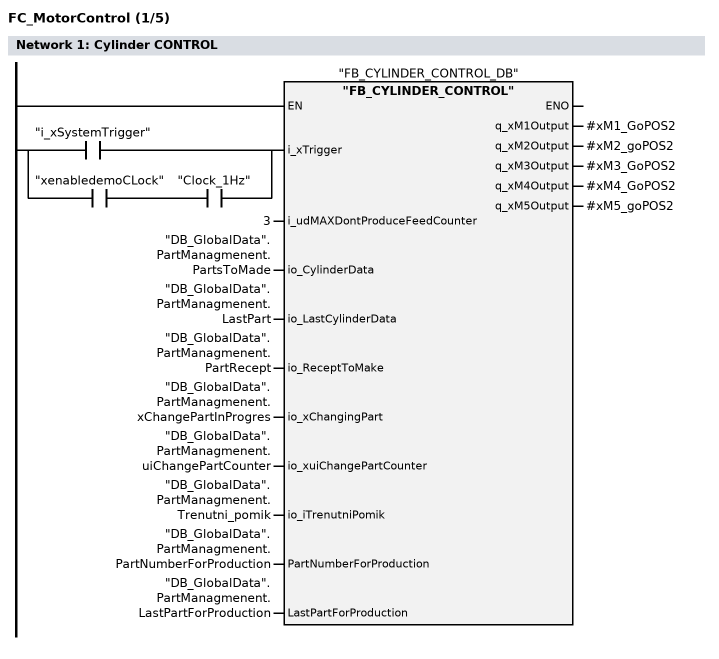
   RUNG wire#powerrail
      "FB_CYLINDER_CONTROL_DB"(i_xTrigger := wire#w1, i_udMAXDontProduceFeedCounter := 3, io_CylinderData := "DB_GlobalData".PartManagmenent.PartsToMade, io_LastCylinderData := "DB_GlobalData".PartManagmenent.LastPart, io_ReceptToMake := "DB_GlobalData".PartManagmenent.PartRecept, io_xChangingPart := "DB_GlobalData".PartManagmenent.xChangePartInProgres, io_xuiChangePartCounter := "DB_GlobalData".PartManagmenent.uiChangePartCounter, io_iTrenutniPomik := "DB_GlobalData".PartManagmenent.Trenutni_pomik, PartNumberForProduction := "DB_GlobalData".PartManagmenent.PartNumberForProduction, LastPartForProduction := "DB_GlobalData".PartManagmenent.LastPartForProduction, q_xM1Output => #xM1_GoPOS2, q_xM2Output => #xM2_goPOS2, q_xM3Output => #xM3_GoPOS2, q_xM4Output => #xM4_GoPOS2, q_xM5Output => #xM5_goPOS2)
   END_RUNG
   RUNG wire#powerrail
      Contact( "i_xSystemTrigger" )
   END_RUNG wire#w1
   RUNG wire#powerrail
      Contact( "xenabledemoCLock" )
      Contact( "Clock_1Hz" )
   END_RUNG wire#w1
   // the same network as SCL:
   "FB_CYLINDER_CONTROL_DB"(i_xTrigger := "i_xSystemTrigger" OR ("xenabledemoCLock" AND "Clock_1Hz"),   // "FB_CYLINDER_CONTROL"
                           i_udMAXDontProduceFeedCounter := 3,
                           io_CylinderData := "DB_GlobalData".PartManagmenent.PartsToMade,
                           io_LastCylinderData := "DB_GlobalData".PartManagmenent.LastPart,
                           io_ReceptToMake := "DB_GlobalData".PartManagmenent.PartRecept,
                           io_xChangingPart := "DB_GlobalData".PartManagmenent.xChangePartInProgres,
                           io_xuiChangePartCounter := "DB_GlobalData".PartManagmenent.uiChangePartCounter,
                           io_iTrenutniPomik := "DB_GlobalData".PartManagmenent.Trenutni_pomik,
                           PartNumberForProduction := "DB_GlobalData".PartManagmenent.PartNumberForProduction,
                           LastPartForProduction := "DB_GlobalData".PartManagmenent.LastPartForProduction,
                           q_xM1Output => #xM1_GoPOS2,
                           q_xM2Output => #xM2_goPOS2,
                           q_xM3Output => #xM3_GoPOS2,
                           q_xM4Output => #xM4_GoPOS2,
                           q_xM5Output => #xM5_goPOS2);
END_REGION

REGION Network 2
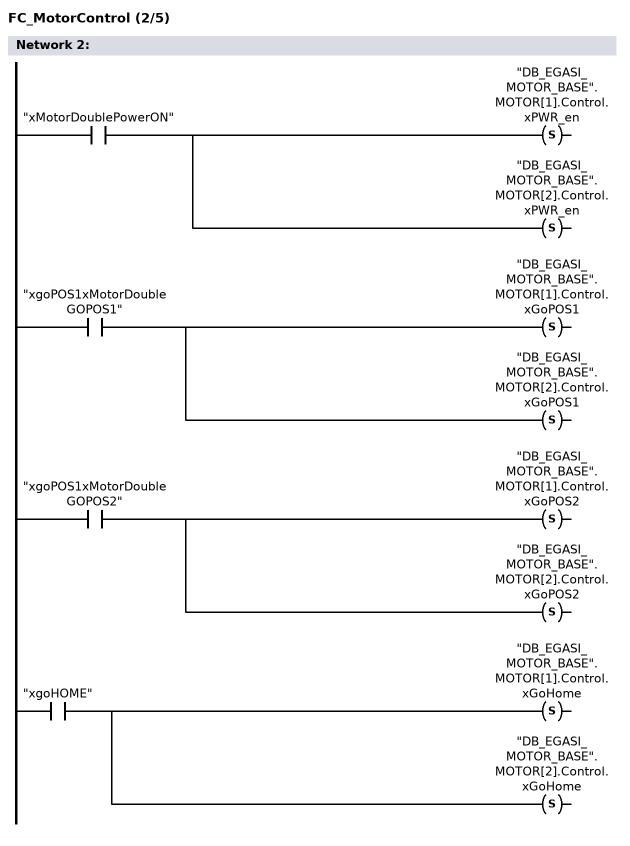
   RUNG wire#powerrail
      Contact( "xMotorDoublePowerON" )
      wire#w1
      S_Coil( "DB_EGASI_MOTOR_BASE".MOTOR[1].Control.xPWR_en )
   END_RUNG
   RUNG wire#w1
      S_Coil( "DB_EGASI_MOTOR_BASE".MOTOR[2].Control.xPWR_en )
   END_RUNG
   RUNG wire#powerrail
      Contact( "xgoPOS1xMotorDoubleGOPOS1" )
      wire#w2
      S_Coil( "DB_EGASI_MOTOR_BASE".MOTOR[1].Control.xGoPOS1 )
   END_RUNG
   RUNG wire#w2
      S_Coil( "DB_EGASI_MOTOR_BASE".MOTOR[2].Control.xGoPOS1 )
   END_RUNG
   RUNG wire#powerrail
      Contact( "xgoPOS1xMotorDoubleGOPOS2" )
      wire#w3
      S_Coil( "DB_EGASI_MOTOR_BASE".MOTOR[1].Control.xGoPOS2 )
   END_RUNG
   RUNG wire#w3
      S_Coil( "DB_EGASI_MOTOR_BASE".MOTOR[2].Control.xGoPOS2 )
   END_RUNG
   RUNG wire#powerrail
      Contact( "xgoHOME" )
      wire#w4
      S_Coil( "DB_EGASI_MOTOR_BASE".MOTOR[1].Control.xGoHome )
   END_RUNG
   RUNG wire#w4
      S_Coil( "DB_EGASI_MOTOR_BASE".MOTOR[2].Control.xGoHome )
   END_RUNG
   // the same network as SCL:
   IF "xMotorDoublePowerON" THEN
       "DB_EGASI_MOTOR_BASE".MOTOR[1].Control.xPWR_en := TRUE;
       "DB_EGASI_MOTOR_BASE".MOTOR[2].Control.xPWR_en := TRUE;
   END_IF;
   IF "xgoPOS1xMotorDoubleGOPOS1" THEN
       "DB_EGASI_MOTOR_BASE".MOTOR[1].Control.xGoPOS1 := TRUE;
       "DB_EGASI_MOTOR_BASE".MOTOR[2].Control.xGoPOS1 := TRUE;
   END_IF;
   IF "xgoPOS1xMotorDoubleGOPOS2" THEN
       "DB_EGASI_MOTOR_BASE".MOTOR[1].Control.xGoPOS2 := TRUE;
       "DB_EGASI_MOTOR_BASE".MOTOR[2].Control.xGoPOS2 := TRUE;
   END_IF;
   IF "xgoHOME" THEN
       "DB_EGASI_MOTOR_BASE".MOTOR[1].Control.xGoHome := TRUE;
       "DB_EGASI_MOTOR_BASE".MOTOR[2].Control.xGoHome := TRUE;
   END_IF;
END_REGION

REGION Network 3: EGASI MOTOR CONTROL
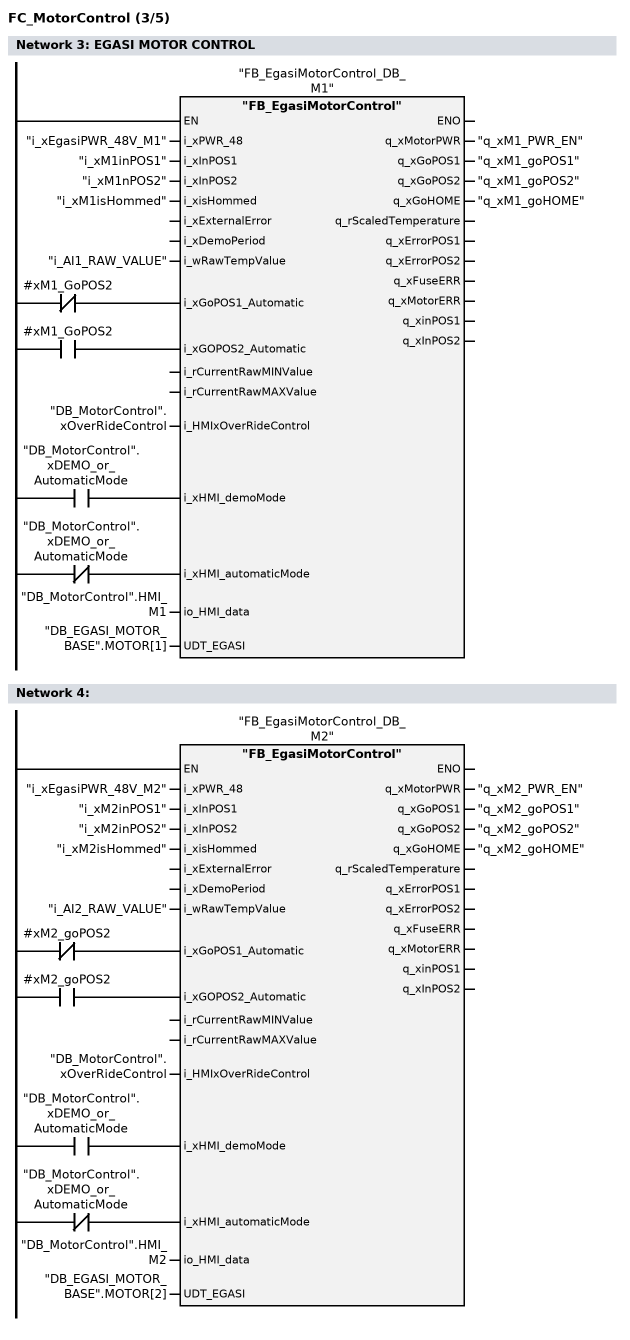
   RUNG wire#powerrail
      "FB_EgasiMotorControl_DB_M1"(i_xGoPOS1_Automatic := wire#w1, i_xGOPOS2_Automatic := wire#w2, i_xHMI_demoMode := wire#w3, i_xHMI_automaticMode := wire#w4, i_xPWR_48 := "i_xEgasiPWR_48V_M1", i_xInPOS1 := "i_xM1inPOS1", i_xInPOS2 := "i_xM1nPOS2", i_xisHommed := "i_xM1isHommed", i_xExternalError :=, i_xDemoPeriod :=, i_wRawTempValue := "i_AI1_RAW_VALUE", i_rCurrentRawMINValue :=, i_rCurrentRawMAXValue :=, i_HMIxOverRideControl := "DB_MotorControl".xOverRideControl, io_HMI_data := "DB_MotorControl".HMI_M1, UDT_EGASI := "DB_EGASI_MOTOR_BASE".MOTOR[1], q_xMotorPWR => "q_xM1_PWR_EN", q_xGoPOS1 => "q_xM1_goPOS1", q_xGoPOS2 => "q_xM1_goPOS2", q_xGoHOME => "q_xM1_goHOME", q_rScaledTemperature =>, q_xErrorPOS1 =>, q_xErrorPOS2 =>, q_xFuseERR =>, q_xMotorERR =>, q_xinPOS1 =>, q_xInPOS2 =>)
   END_RUNG
   RUNG wire#powerrail
      I_Contact( #xM1_GoPOS2 )
   END_RUNG wire#w1
   RUNG wire#powerrail
      Contact( #xM1_GoPOS2 )
   END_RUNG wire#w2
   RUNG wire#powerrail
      Contact( "DB_MotorControl".xDEMO_or_AutomaticMode )
   END_RUNG wire#w3
   RUNG wire#powerrail
      I_Contact( "DB_MotorControl".xDEMO_or_AutomaticMode )
   END_RUNG wire#w4
   // the same network as SCL:
   "FB_EgasiMotorControl_DB_M1"(i_xPWR_48 := "i_xEgasiPWR_48V_M1",   // "FB_EgasiMotorControl"
                           i_xInPOS1 := "i_xM1inPOS1",
                           i_xInPOS2 := "i_xM1nPOS2",
                           i_xisHommed := "i_xM1isHommed",
                           i_wRawTempValue := "i_AI1_RAW_VALUE",
                           i_xGoPOS1_Automatic := NOT #xM1_GoPOS2,
                           i_xGOPOS2_Automatic := #xM1_GoPOS2,
                           i_HMIxOverRideControl := "DB_MotorControl".xOverRideControl,
                           i_xHMI_demoMode := "DB_MotorControl".xDEMO_or_AutomaticMode,
                           i_xHMI_automaticMode := NOT "DB_MotorControl".xDEMO_or_AutomaticMode,
                           io_HMI_data := "DB_MotorControl".HMI_M1,
                           UDT_EGASI := "DB_EGASI_MOTOR_BASE".MOTOR[1],
                           q_xMotorPWR => "q_xM1_PWR_EN",
                           q_xGoPOS1 => "q_xM1_goPOS1",
                           q_xGoPOS2 => "q_xM1_goPOS2",
                           q_xGoHOME => "q_xM1_goHOME");
END_REGION

REGION Network 4
   RUNG wire#powerrail
      "FB_EgasiMotorControl_DB_M2"(i_xGoPOS1_Automatic := wire#w1, i_xGOPOS2_Automatic := wire#w2, i_xHMI_demoMode := wire#w3, i_xHMI_automaticMode := wire#w4, i_xPWR_48 := "i_xEgasiPWR_48V_M2", i_xInPOS1 := "i_xM2inPOS1", i_xInPOS2 := "i_xM2inPOS2", i_xisHommed := "i_xM2isHommed", i_xExternalError :=, i_xDemoPeriod :=, i_wRawTempValue := "i_AI2_RAW_VALUE", i_rCurrentRawMINValue :=, i_rCurrentRawMAXValue :=, i_HMIxOverRideControl := "DB_MotorControl".xOverRideControl, io_HMI_data := "DB_MotorControl".HMI_M2, UDT_EGASI := "DB_EGASI_MOTOR_BASE".MOTOR[2], q_xMotorPWR => "q_xM2_PWR_EN", q_xGoPOS1 => "q_xM2_goPOS1", q_xGoPOS2 => "q_xM2_goPOS2", q_xGoHOME => "q_xM2_goHOME", q_rScaledTemperature =>, q_xErrorPOS1 =>, q_xErrorPOS2 =>, q_xFuseERR =>, q_xMotorERR =>, q_xinPOS1 =>, q_xInPOS2 =>)
   END_RUNG
   RUNG wire#powerrail
      I_Contact( #xM2_goPOS2 )
   END_RUNG wire#w1
   RUNG wire#powerrail
      Contact( #xM2_goPOS2 )
   END_RUNG wire#w2
   RUNG wire#powerrail
      Contact( "DB_MotorControl".xDEMO_or_AutomaticMode )
   END_RUNG wire#w3
   RUNG wire#powerrail
      I_Contact( "DB_MotorControl".xDEMO_or_AutomaticMode )
   END_RUNG wire#w4
   // the same network as SCL:
   "FB_EgasiMotorControl_DB_M2"(i_xPWR_48 := "i_xEgasiPWR_48V_M2",   // "FB_EgasiMotorControl"
                           i_xInPOS1 := "i_xM2inPOS1",
                           i_xInPOS2 := "i_xM2inPOS2",
                           i_xisHommed := "i_xM2isHommed",
                           i_wRawTempValue := "i_AI2_RAW_VALUE",
                           i_xGoPOS1_Automatic := NOT #xM2_goPOS2,
                           i_xGOPOS2_Automatic := #xM2_goPOS2,
                           i_HMIxOverRideControl := "DB_MotorControl".xOverRideControl,
                           i_xHMI_demoMode := "DB_MotorControl".xDEMO_or_AutomaticMode,
                           i_xHMI_automaticMode := NOT "DB_MotorControl".xDEMO_or_AutomaticMode,
                           io_HMI_data := "DB_MotorControl".HMI_M2,
                           UDT_EGASI := "DB_EGASI_MOTOR_BASE".MOTOR[2],
                           q_xMotorPWR => "q_xM2_PWR_EN",
                           q_xGoPOS1 => "q_xM2_goPOS1",
                           q_xGoPOS2 => "q_xM2_goPOS2",
                           q_xGoHOME => "q_xM2_goHOME");
END_REGION

REGION Network 5
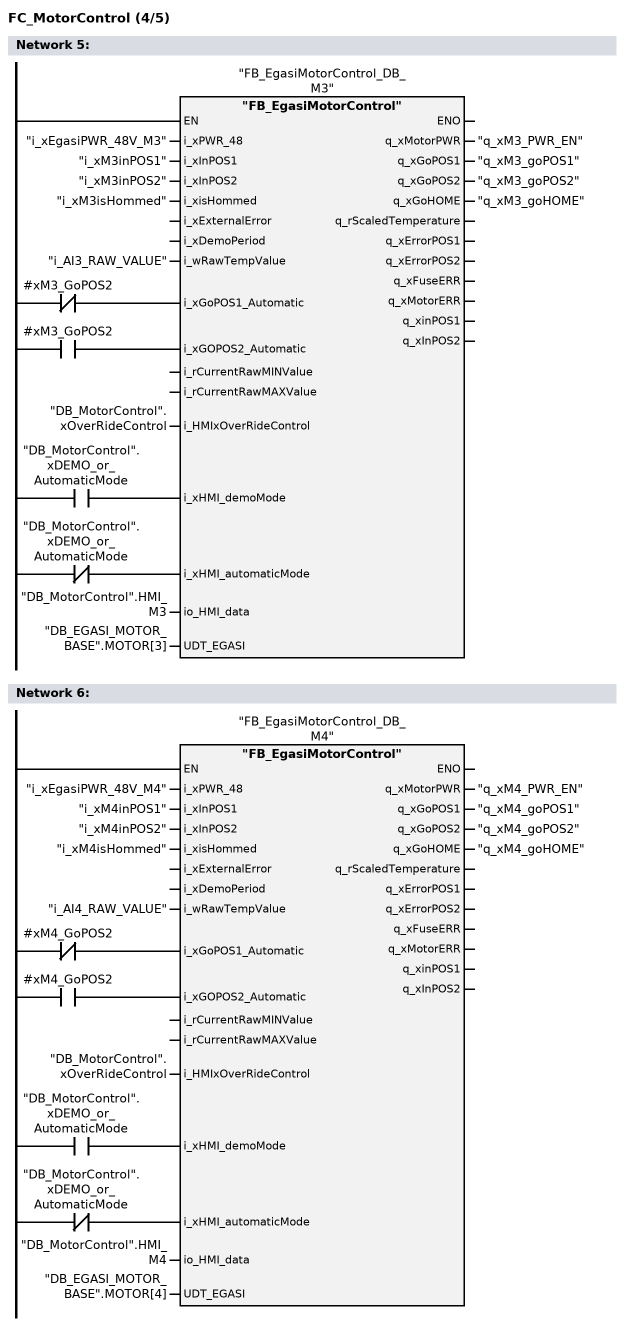
   RUNG wire#powerrail
      "FB_EgasiMotorControl_DB_M3"(i_xGoPOS1_Automatic := wire#w1, i_xGOPOS2_Automatic := wire#w2, i_xHMI_demoMode := wire#w3, i_xHMI_automaticMode := wire#w4, i_xPWR_48 := "i_xEgasiPWR_48V_M3", i_xInPOS1 := "i_xM3inPOS1", i_xInPOS2 := "i_xM3inPOS2", i_xisHommed := "i_xM3isHommed", i_xExternalError :=, i_xDemoPeriod :=, i_wRawTempValue := "i_AI3_RAW_VALUE", i_rCurrentRawMINValue :=, i_rCurrentRawMAXValue :=, i_HMIxOverRideControl := "DB_MotorControl".xOverRideControl, io_HMI_data := "DB_MotorControl".HMI_M3, UDT_EGASI := "DB_EGASI_MOTOR_BASE".MOTOR[3], q_xMotorPWR => "q_xM3_PWR_EN", q_xGoPOS1 => "q_xM3_goPOS1", q_xGoPOS2 => "q_xM3_goPOS2", q_xGoHOME => "q_xM3_goHOME", q_rScaledTemperature =>, q_xErrorPOS1 =>, q_xErrorPOS2 =>, q_xFuseERR =>, q_xMotorERR =>, q_xinPOS1 =>, q_xInPOS2 =>)
   END_RUNG
   RUNG wire#powerrail
      I_Contact( #xM3_GoPOS2 )
   END_RUNG wire#w1
   RUNG wire#powerrail
      Contact( #xM3_GoPOS2 )
   END_RUNG wire#w2
   RUNG wire#powerrail
      Contact( "DB_MotorControl".xDEMO_or_AutomaticMode )
   END_RUNG wire#w3
   RUNG wire#powerrail
      I_Contact( "DB_MotorControl".xDEMO_or_AutomaticMode )
   END_RUNG wire#w4
   // the same network as SCL:
   "FB_EgasiMotorControl_DB_M3"(i_xPWR_48 := "i_xEgasiPWR_48V_M3",   // "FB_EgasiMotorControl"
                           i_xInPOS1 := "i_xM3inPOS1",
                           i_xInPOS2 := "i_xM3inPOS2",
                           i_xisHommed := "i_xM3isHommed",
                           i_wRawTempValue := "i_AI3_RAW_VALUE",
                           i_xGoPOS1_Automatic := NOT #xM3_GoPOS2,
                           i_xGOPOS2_Automatic := #xM3_GoPOS2,
                           i_HMIxOverRideControl := "DB_MotorControl".xOverRideControl,
                           i_xHMI_demoMode := "DB_MotorControl".xDEMO_or_AutomaticMode,
                           i_xHMI_automaticMode := NOT "DB_MotorControl".xDEMO_or_AutomaticMode,
                           io_HMI_data := "DB_MotorControl".HMI_M3,
                           UDT_EGASI := "DB_EGASI_MOTOR_BASE".MOTOR[3],
                           q_xMotorPWR => "q_xM3_PWR_EN",
                           q_xGoPOS1 => "q_xM3_goPOS1",
                           q_xGoPOS2 => "q_xM3_goPOS2",
                           q_xGoHOME => "q_xM3_goHOME");
END_REGION

REGION Network 6
   RUNG wire#powerrail
      "FB_EgasiMotorControl_DB_M4"(i_xGoPOS1_Automatic := wire#w1, i_xGOPOS2_Automatic := wire#w2, i_xHMI_demoMode := wire#w3, i_xHMI_automaticMode := wire#w4, i_xPWR_48 := "i_xEgasiPWR_48V_M4", i_xInPOS1 := "i_xM4inPOS1", i_xInPOS2 := "i_xM4inPOS2", i_xisHommed := "i_xM4isHommed", i_xExternalError :=, i_xDemoPeriod :=, i_wRawTempValue := "i_AI4_RAW_VALUE", i_rCurrentRawMINValue :=, i_rCurrentRawMAXValue :=, i_HMIxOverRideControl := "DB_MotorControl".xOverRideControl, io_HMI_data := "DB_MotorControl".HMI_M4, UDT_EGASI := "DB_EGASI_MOTOR_BASE".MOTOR[4], q_xMotorPWR => "q_xM4_PWR_EN", q_xGoPOS1 => "q_xM4_goPOS1", q_xGoPOS2 => "q_xM4_goPOS2", q_xGoHOME => "q_xM4_goHOME", q_rScaledTemperature =>, q_xErrorPOS1 =>, q_xErrorPOS2 =>, q_xFuseERR =>, q_xMotorERR =>, q_xinPOS1 =>, q_xInPOS2 =>)
   END_RUNG
   RUNG wire#powerrail
      I_Contact( #xM4_GoPOS2 )
   END_RUNG wire#w1
   RUNG wire#powerrail
      Contact( #xM4_GoPOS2 )
   END_RUNG wire#w2
   RUNG wire#powerrail
      Contact( "DB_MotorControl".xDEMO_or_AutomaticMode )
   END_RUNG wire#w3
   RUNG wire#powerrail
      I_Contact( "DB_MotorControl".xDEMO_or_AutomaticMode )
   END_RUNG wire#w4
   // the same network as SCL:
   "FB_EgasiMotorControl_DB_M4"(i_xPWR_48 := "i_xEgasiPWR_48V_M4",   // "FB_EgasiMotorControl"
                           i_xInPOS1 := "i_xM4inPOS1",
                           i_xInPOS2 := "i_xM4inPOS2",
                           i_xisHommed := "i_xM4isHommed",
                           i_wRawTempValue := "i_AI4_RAW_VALUE",
                           i_xGoPOS1_Automatic := NOT #xM4_GoPOS2,
                           i_xGOPOS2_Automatic := #xM4_GoPOS2,
                           i_HMIxOverRideControl := "DB_MotorControl".xOverRideControl,
                           i_xHMI_demoMode := "DB_MotorControl".xDEMO_or_AutomaticMode,
                           i_xHMI_automaticMode := NOT "DB_MotorControl".xDEMO_or_AutomaticMode,
                           io_HMI_data := "DB_MotorControl".HMI_M4,
                           UDT_EGASI := "DB_EGASI_MOTOR_BASE".MOTOR[4],
                           q_xMotorPWR => "q_xM4_PWR_EN",
                           q_xGoPOS1 => "q_xM4_goPOS1",
                           q_xGoPOS2 => "q_xM4_goPOS2",
                           q_xGoHOME => "q_xM4_goHOME");
END_REGION

REGION Network 7
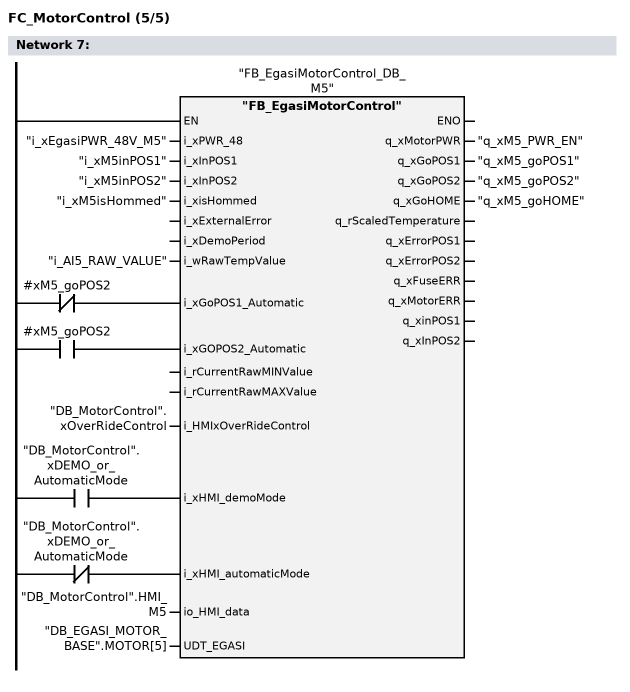
   RUNG wire#powerrail
      "FB_EgasiMotorControl_DB_M5"(i_xGoPOS1_Automatic := wire#w1, i_xGOPOS2_Automatic := wire#w2, i_xHMI_demoMode := wire#w3, i_xHMI_automaticMode := wire#w4, i_xPWR_48 := "i_xEgasiPWR_48V_M5", i_xInPOS1 := "i_xM5inPOS1", i_xInPOS2 := "i_xM5inPOS2", i_xisHommed := "i_xM5isHommed", i_xExternalError :=, i_xDemoPeriod :=, i_wRawTempValue := "i_AI5_RAW_VALUE", i_rCurrentRawMINValue :=, i_rCurrentRawMAXValue :=, i_HMIxOverRideControl := "DB_MotorControl".xOverRideControl, io_HMI_data := "DB_MotorControl".HMI_M5, UDT_EGASI := "DB_EGASI_MOTOR_BASE".MOTOR[5], q_xMotorPWR => "q_xM5_PWR_EN", q_xGoPOS1 => "q_xM5_goPOS1", q_xGoPOS2 => "q_xM5_goPOS2", q_xGoHOME => "q_xM5_goHOME", q_rScaledTemperature =>, q_xErrorPOS1 =>, q_xErrorPOS2 =>, q_xFuseERR =>, q_xMotorERR =>, q_xinPOS1 =>, q_xInPOS2 =>)
   END_RUNG
   RUNG wire#powerrail
      I_Contact( #xM5_goPOS2 )
   END_RUNG wire#w1
   RUNG wire#powerrail
      Contact( #xM5_goPOS2 )
   END_RUNG wire#w2
   RUNG wire#powerrail
      Contact( "DB_MotorControl".xDEMO_or_AutomaticMode )
   END_RUNG wire#w3
   RUNG wire#powerrail
      I_Contact( "DB_MotorControl".xDEMO_or_AutomaticMode )
   END_RUNG wire#w4
   // the same network as SCL:
   "FB_EgasiMotorControl_DB_M5"(i_xPWR_48 := "i_xEgasiPWR_48V_M5",   // "FB_EgasiMotorControl"
                           i_xInPOS1 := "i_xM5inPOS1",
                           i_xInPOS2 := "i_xM5inPOS2",
                           i_xisHommed := "i_xM5isHommed",
                           i_wRawTempValue := "i_AI5_RAW_VALUE",
                           i_xGoPOS1_Automatic := NOT #xM5_goPOS2,
                           i_xGOPOS2_Automatic := #xM5_goPOS2,
                           i_HMIxOverRideControl := "DB_MotorControl".xOverRideControl,
                           i_xHMI_demoMode := "DB_MotorControl".xDEMO_or_AutomaticMode,
                           i_xHMI_automaticMode := NOT "DB_MotorControl".xDEMO_or_AutomaticMode,
                           io_HMI_data := "DB_MotorControl".HMI_M5,
                           UDT_EGASI := "DB_EGASI_MOTOR_BASE".MOTOR[5],
                           q_xMotorPWR => "q_xM5_PWR_EN",
                           q_xGoPOS1 => "q_xM5_goPOS1",
                           q_xGoPOS2 => "q_xM5_goPOS2",
                           q_xGoHOME => "q_xM5_goHOME");
END_REGION
END_FUNCTION

FUNCTION "FC_PARTMANAGE" : Void   // FC12, LAD
{ S7_Optimized_Access := 'TRUE' }
VERSION : 0.1
   VAR_TEMP   // added for the SCL form of the ladder/FBD networks
      _w1 : Bool;
   END_VAR
BEGIN

REGION Network 2: COPY DATA FROM BASE TO DB for Cylinder control
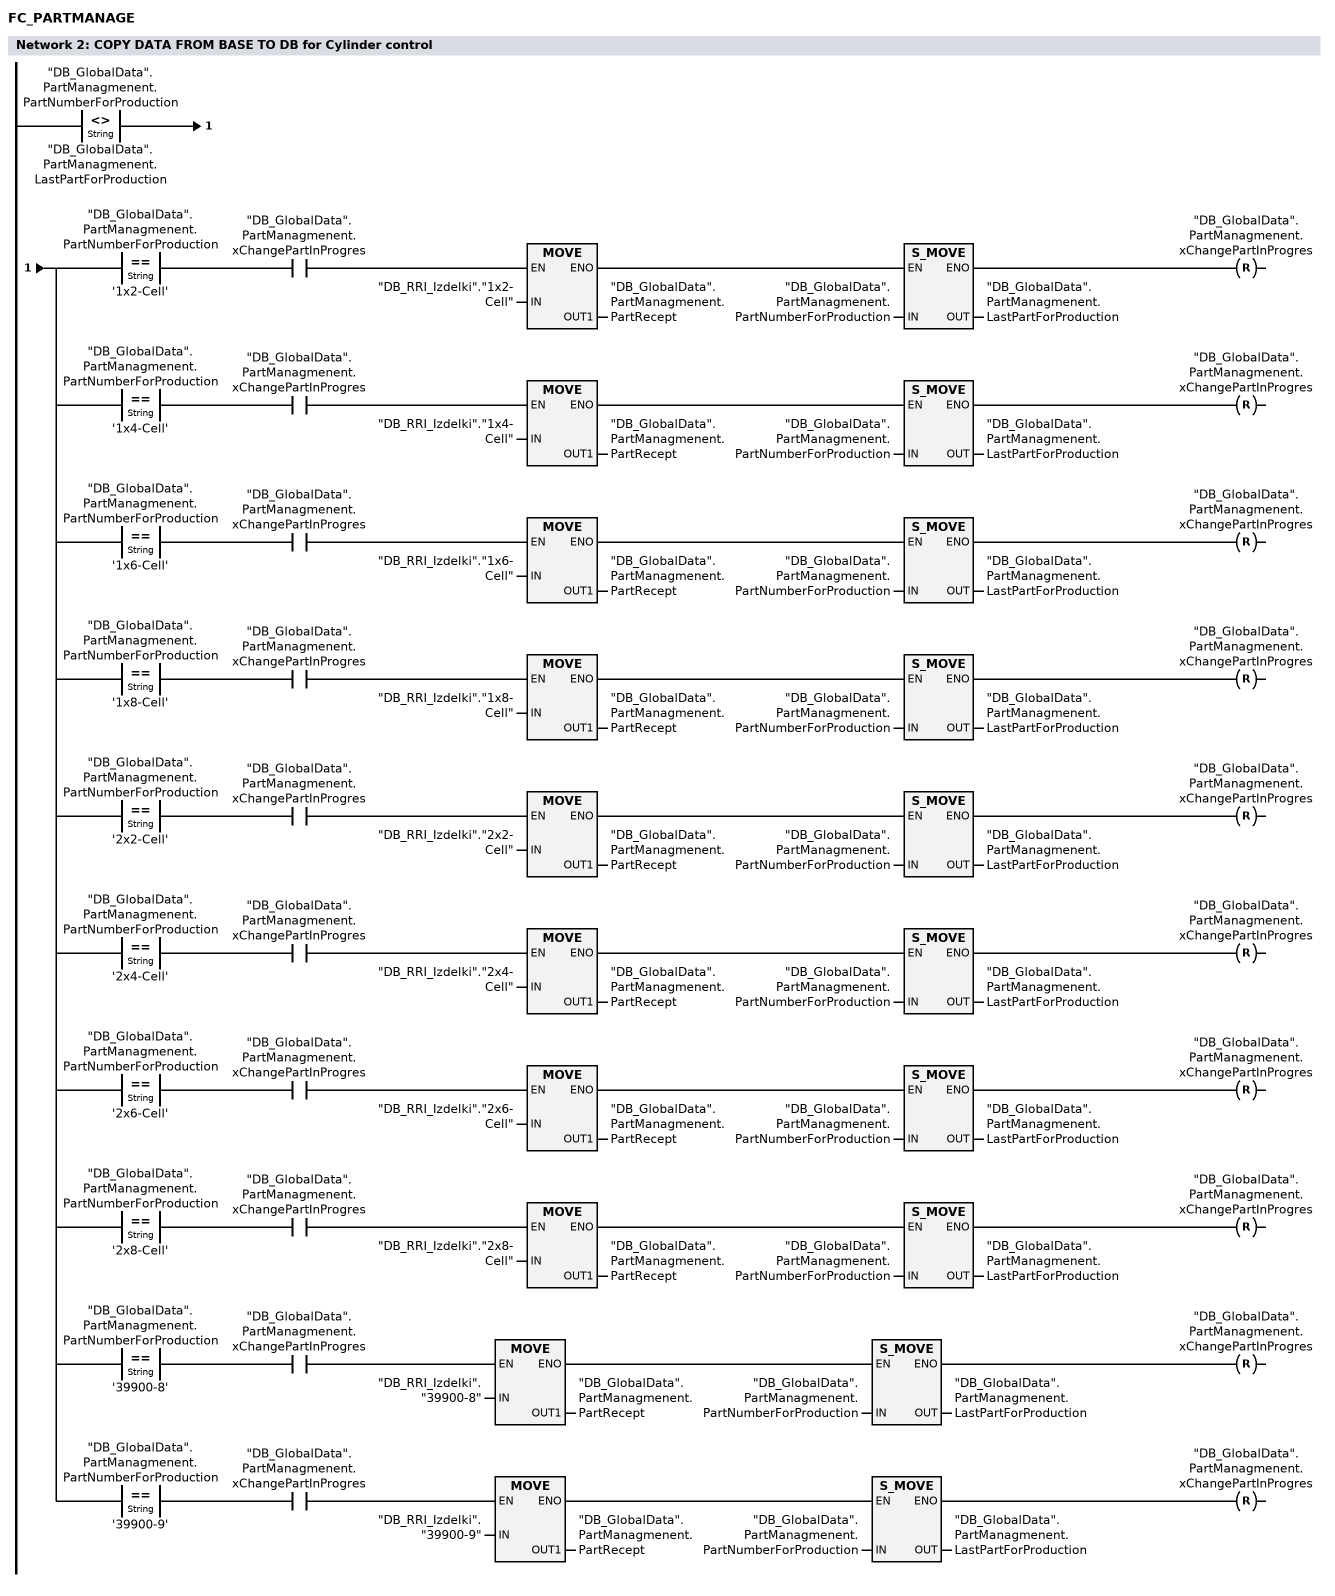
   RUNG wire#powerrail
      { S7_Templates := "SrcType := String" } NE_Contact(in1 := "DB_GlobalData".PartManagmenent.PartNumberForProduction, in2 := "DB_GlobalData".PartManagmenent.LastPartForProduction)
      wire#w1
      { S7_Templates := "SrcType := String" } EQ_Contact(in1 := "DB_GlobalData".PartManagmenent.PartNumberForProduction, in2 := '1x2-Cell')
      Contact( "DB_GlobalData".PartManagmenent.xChangePartInProgres )
      Move(in := "DB_RRI_Izdelki"."1x2-Cell", out1 => "DB_GlobalData".PartManagmenent.PartRecept)
      S_Move(in := "DB_GlobalData".PartManagmenent.PartNumberForProduction, out => "DB_GlobalData".PartManagmenent.LastPartForProduction)
      R_Coil( "DB_GlobalData".PartManagmenent.xChangePartInProgres )
   END_RUNG
   RUNG wire#w1
      { S7_Templates := "SrcType := String" } EQ_Contact(in1 := "DB_GlobalData".PartManagmenent.PartNumberForProduction, in2 := '1x4-Cell')
      Contact( "DB_GlobalData".PartManagmenent.xChangePartInProgres )
      Move(in := "DB_RRI_Izdelki"."1x4-Cell", out1 => "DB_GlobalData".PartManagmenent.PartRecept)
      S_Move(in := "DB_GlobalData".PartManagmenent.PartNumberForProduction, out => "DB_GlobalData".PartManagmenent.LastPartForProduction)
      R_Coil( "DB_GlobalData".PartManagmenent.xChangePartInProgres )
   END_RUNG
   RUNG wire#w1
      { S7_Templates := "SrcType := String" } EQ_Contact(in1 := "DB_GlobalData".PartManagmenent.PartNumberForProduction, in2 := '1x6-Cell')
      Contact( "DB_GlobalData".PartManagmenent.xChangePartInProgres )
      Move(in := "DB_RRI_Izdelki"."1x6-Cell", out1 => "DB_GlobalData".PartManagmenent.PartRecept)
      S_Move(in := "DB_GlobalData".PartManagmenent.PartNumberForProduction, out => "DB_GlobalData".PartManagmenent.LastPartForProduction)
      R_Coil( "DB_GlobalData".PartManagmenent.xChangePartInProgres )
   END_RUNG
   RUNG wire#w1
      { S7_Templates := "SrcType := String" } EQ_Contact(in1 := "DB_GlobalData".PartManagmenent.PartNumberForProduction, in2 := '1x8-Cell')
      Contact( "DB_GlobalData".PartManagmenent.xChangePartInProgres )
      Move(in := "DB_RRI_Izdelki"."1x8-Cell", out1 => "DB_GlobalData".PartManagmenent.PartRecept)
      S_Move(in := "DB_GlobalData".PartManagmenent.PartNumberForProduction, out => "DB_GlobalData".PartManagmenent.LastPartForProduction)
      R_Coil( "DB_GlobalData".PartManagmenent.xChangePartInProgres )
   END_RUNG
   RUNG wire#w1
      { S7_Templates := "SrcType := String" } EQ_Contact(in1 := "DB_GlobalData".PartManagmenent.PartNumberForProduction, in2 := '2x2-Cell')
      Contact( "DB_GlobalData".PartManagmenent.xChangePartInProgres )
      Move(in := "DB_RRI_Izdelki"."2x2-Cell", out1 => "DB_GlobalData".PartManagmenent.PartRecept)
      S_Move(in := "DB_GlobalData".PartManagmenent.PartNumberForProduction, out => "DB_GlobalData".PartManagmenent.LastPartForProduction)
      R_Coil( "DB_GlobalData".PartManagmenent.xChangePartInProgres )
   END_RUNG
   RUNG wire#w1
      { S7_Templates := "SrcType := String" } EQ_Contact(in1 := "DB_GlobalData".PartManagmenent.PartNumberForProduction, in2 := '2x4-Cell')
      Contact( "DB_GlobalData".PartManagmenent.xChangePartInProgres )
      Move(in := "DB_RRI_Izdelki"."2x4-Cell", out1 => "DB_GlobalData".PartManagmenent.PartRecept)
      S_Move(in := "DB_GlobalData".PartManagmenent.PartNumberForProduction, out => "DB_GlobalData".PartManagmenent.LastPartForProduction)
      R_Coil( "DB_GlobalData".PartManagmenent.xChangePartInProgres )
   END_RUNG
   RUNG wire#w1
      { S7_Templates := "SrcType := String" } EQ_Contact(in1 := "DB_GlobalData".PartManagmenent.PartNumberForProduction, in2 := '2x6-Cell')
      Contact( "DB_GlobalData".PartManagmenent.xChangePartInProgres )
      Move(in := "DB_RRI_Izdelki"."2x6-Cell", out1 => "DB_GlobalData".PartManagmenent.PartRecept)
      S_Move(in := "DB_GlobalData".PartManagmenent.PartNumberForProduction, out => "DB_GlobalData".PartManagmenent.LastPartForProduction)
      R_Coil( "DB_GlobalData".PartManagmenent.xChangePartInProgres )
   END_RUNG
   RUNG wire#w1
      { S7_Templates := "SrcType := String" } EQ_Contact(in1 := "DB_GlobalData".PartManagmenent.PartNumberForProduction, in2 := '2x8-Cell')
      Contact( "DB_GlobalData".PartManagmenent.xChangePartInProgres )
      Move(in := "DB_RRI_Izdelki"."2x8-Cell", out1 => "DB_GlobalData".PartManagmenent.PartRecept)
      S_Move(in := "DB_GlobalData".PartManagmenent.PartNumberForProduction, out => "DB_GlobalData".PartManagmenent.LastPartForProduction)
      R_Coil( "DB_GlobalData".PartManagmenent.xChangePartInProgres )
   END_RUNG
   RUNG wire#w1
      { S7_Templates := "SrcType := String" } EQ_Contact(in1 := "DB_GlobalData".PartManagmenent.PartNumberForProduction, in2 := '39900-8')
      Contact( "DB_GlobalData".PartManagmenent.xChangePartInProgres )
      Move(in := "DB_RRI_Izdelki"."39900-8", out1 => "DB_GlobalData".PartManagmenent.PartRecept)
      S_Move(in := "DB_GlobalData".PartManagmenent.PartNumberForProduction, out => "DB_GlobalData".PartManagmenent.LastPartForProduction)
      R_Coil( "DB_GlobalData".PartManagmenent.xChangePartInProgres )
   END_RUNG
   RUNG wire#w1
      { S7_Templates := "SrcType := String" } EQ_Contact(in1 := "DB_GlobalData".PartManagmenent.PartNumberForProduction, in2 := '39900-9')
      Contact( "DB_GlobalData".PartManagmenent.xChangePartInProgres )
      Move(in := "DB_RRI_Izdelki"."39900-9", out1 => "DB_GlobalData".PartManagmenent.PartRecept)
      S_Move(in := "DB_GlobalData".PartManagmenent.PartNumberForProduction, out => "DB_GlobalData".PartManagmenent.LastPartForProduction)
      R_Coil( "DB_GlobalData".PartManagmenent.xChangePartInProgres )
   END_RUNG
   // the same network as SCL:
   #_w1 := "DB_GlobalData".PartManagmenent.PartNumberForProduction <> "DB_GlobalData".PartManagmenent.LastPartForProduction;
   IF #_w1 AND ("DB_GlobalData".PartManagmenent.PartNumberForProduction = '1x2-Cell') AND "DB_GlobalData".PartManagmenent.xChangePartInProgres THEN
       "DB_GlobalData".PartManagmenent.PartRecept := "DB_RRI_Izdelki"."1x2-Cell";
       "DB_GlobalData".PartManagmenent.LastPartForProduction := "DB_GlobalData".PartManagmenent.PartNumberForProduction;
       "DB_GlobalData".PartManagmenent.xChangePartInProgres := FALSE;
   END_IF;
   IF #_w1 AND ("DB_GlobalData".PartManagmenent.PartNumberForProduction = '1x4-Cell') AND "DB_GlobalData".PartManagmenent.xChangePartInProgres THEN
       "DB_GlobalData".PartManagmenent.PartRecept := "DB_RRI_Izdelki"."1x4-Cell";
       "DB_GlobalData".PartManagmenent.LastPartForProduction := "DB_GlobalData".PartManagmenent.PartNumberForProduction;
       "DB_GlobalData".PartManagmenent.xChangePartInProgres := FALSE;
   END_IF;
   IF #_w1 AND ("DB_GlobalData".PartManagmenent.PartNumberForProduction = '1x6-Cell') AND "DB_GlobalData".PartManagmenent.xChangePartInProgres THEN
       "DB_GlobalData".PartManagmenent.PartRecept := "DB_RRI_Izdelki"."1x6-Cell";
       "DB_GlobalData".PartManagmenent.LastPartForProduction := "DB_GlobalData".PartManagmenent.PartNumberForProduction;
       "DB_GlobalData".PartManagmenent.xChangePartInProgres := FALSE;
   END_IF;
   IF #_w1 AND ("DB_GlobalData".PartManagmenent.PartNumberForProduction = '1x8-Cell') AND "DB_GlobalData".PartManagmenent.xChangePartInProgres THEN
       "DB_GlobalData".PartManagmenent.PartRecept := "DB_RRI_Izdelki"."1x8-Cell";
       "DB_GlobalData".PartManagmenent.LastPartForProduction := "DB_GlobalData".PartManagmenent.PartNumberForProduction;
       "DB_GlobalData".PartManagmenent.xChangePartInProgres := FALSE;
   END_IF;
   IF #_w1 AND ("DB_GlobalData".PartManagmenent.PartNumberForProduction = '2x2-Cell') AND "DB_GlobalData".PartManagmenent.xChangePartInProgres THEN
       "DB_GlobalData".PartManagmenent.PartRecept := "DB_RRI_Izdelki"."2x2-Cell";
       "DB_GlobalData".PartManagmenent.LastPartForProduction := "DB_GlobalData".PartManagmenent.PartNumberForProduction;
       "DB_GlobalData".PartManagmenent.xChangePartInProgres := FALSE;
   END_IF;
   IF #_w1 AND ("DB_GlobalData".PartManagmenent.PartNumberForProduction = '2x4-Cell') AND "DB_GlobalData".PartManagmenent.xChangePartInProgres THEN
       "DB_GlobalData".PartManagmenent.PartRecept := "DB_RRI_Izdelki"."2x4-Cell";
       "DB_GlobalData".PartManagmenent.LastPartForProduction := "DB_GlobalData".PartManagmenent.PartNumberForProduction;
       "DB_GlobalData".PartManagmenent.xChangePartInProgres := FALSE;
   END_IF;
   IF #_w1 AND ("DB_GlobalData".PartManagmenent.PartNumberForProduction = '2x6-Cell') AND "DB_GlobalData".PartManagmenent.xChangePartInProgres THEN
       "DB_GlobalData".PartManagmenent.PartRecept := "DB_RRI_Izdelki"."2x6-Cell";
       "DB_GlobalData".PartManagmenent.LastPartForProduction := "DB_GlobalData".PartManagmenent.PartNumberForProduction;
       "DB_GlobalData".PartManagmenent.xChangePartInProgres := FALSE;
   END_IF;
   IF #_w1 AND ("DB_GlobalData".PartManagmenent.PartNumberForProduction = '2x8-Cell') AND "DB_GlobalData".PartManagmenent.xChangePartInProgres THEN
       "DB_GlobalData".PartManagmenent.PartRecept := "DB_RRI_Izdelki"."2x8-Cell";
       "DB_GlobalData".PartManagmenent.LastPartForProduction := "DB_GlobalData".PartManagmenent.PartNumberForProduction;
       "DB_GlobalData".PartManagmenent.xChangePartInProgres := FALSE;
   END_IF;
   IF #_w1 AND ("DB_GlobalData".PartManagmenent.PartNumberForProduction = '39900-8') AND "DB_GlobalData".PartManagmenent.xChangePartInProgres THEN
       "DB_GlobalData".PartManagmenent.PartRecept := "DB_RRI_Izdelki"."39900-8";
       "DB_GlobalData".PartManagmenent.LastPartForProduction := "DB_GlobalData".PartManagmenent.PartNumberForProduction;
       "DB_GlobalData".PartManagmenent.xChangePartInProgres := FALSE;
   END_IF;
   IF #_w1 AND ("DB_GlobalData".PartManagmenent.PartNumberForProduction = '39900-9') AND "DB_GlobalData".PartManagmenent.xChangePartInProgres THEN
       "DB_GlobalData".PartManagmenent.PartRecept := "DB_RRI_Izdelki"."39900-9";
       "DB_GlobalData".PartManagmenent.LastPartForProduction := "DB_GlobalData".PartManagmenent.PartNumberForProduction;
       "DB_GlobalData".PartManagmenent.xChangePartInProgres := FALSE;
   END_IF;
END_REGION
